ADD_ON_INSTRUCTION GP_HeadPositionDefined   (* revision 1.0 *)
// To be called before invertion data
VAR_IN_OUT
   In_ConvoyData : UDT_Convoy_SL; {required}
END_VAR
VAR_INPUT
   In_dConveyorLenght : DINT; {access None, required}   // Conveyor below [mm/100]
   In_dConveyorWidth : DINT; {access None, required}   // Conveyor below [mm/100]
   In_dInLitePos : DINT; {access None, required}   // Position input lite - Left to Right line flow(0=AX; 1=XA)
   In_dOutDirection : DINT; {required}   // Direction of lateral flow (0=Left; 1=Right; 2=CW(rotation); 3=CCW(rotation))
   In_dOutLitePos : DINT; {access None, required}   // Position output lite - Left to Right line flow(0=AX; 1=XA)
END_VAR
VAR_OUTPUT
   Out_dHeadPosition : DINT; {access Read Only, required}   // New head position [mm/100]
END_VAR
VAR
   TMP_idxCap : DINT; {access None}
   TMP_IdxLite : DINT; {access None}
   TMP_MaxCap : DINT; {access None}
   TMP_MaxLite : DINT; {access None}
   TMP_d : DINT; {access None}
   TMP_LiteHeadReference : DINT; {access None}   // New convoy lite head [mm/100]
END_VAR

ROUTINE Logic   (* structured text *)
   ////////////////////////////////////////////////////////////
   //   Copyright (c)  <Key Automation srl>
   //------------------------------------------------------------
   //   Routine: GP_HeadPositionDefined - Logic
   //   Author: Gerto\admin
   //   Created: 2020-02-05
   //------------------------------------------------------------
   //   Description:
   //
   //
   //   History:
   //
   ////////////////////////////////////////////////////////////
   
   //Dimension array
   Size(In_ConvoyData.rgtCap,0,TMP_MaxCap);
   size(In_ConvoyData.rgtCap[0].rgtLite,0,TMP_MaxLite);
   
   //Find lite of reference
   
   // The smallest LitesHead (Barycenter Lite - 1/2 width lite)
   if 	(In_dOutDirection = 0 and In_dInLitePos = 0 and In_dOutLitePos = 0) or
   	(In_dOutDirection = 0 and In_dInLitePos = 0 and In_dOutLitePos = 1) or
   	(In_dOutDirection = 1 and In_dInLitePos = 1 and In_dOutLitePos = 0) or
   	(In_dOutDirection = 1 and In_dInLitePos = 1 and In_dOutLitePos = 1) or
   	(In_dOutDirection = 2 and In_dInLitePos = 0 and In_dOutLitePos = 0) or
   	(In_dOutDirection = 3 and In_dInLitePos = 1 and In_dOutLitePos = 1) then
   	TMP_LiteHeadReference := In_dConveyorWidth;
   	For TMP_idxCap := 0 to TMP_MaxCap-1 by 1 do
   		for TMP_IdxLite := 0 to TMP_MaxLite-1 by 1 do
   			if In_ConvoyData.rgtCap[TMP_idxCap].rgtLite[TMP_IdxLite].dID <> 0 and (In_ConvoyData.rgtCap[TMP_idxCap].rgtLite[TMP_IdxLite].dBarycenter_cmm - In_ConvoyData.rgtCap[TMP_idxCap].rgtLite[TMP_IdxLite].dWidth_cmm/2) < TMP_LiteHeadReference then
   				TMP_LiteHeadReference := In_ConvoyData.rgtCap[TMP_idxCap].rgtLite[TMP_IdxLite].dBarycenter_cmm - In_ConvoyData.rgtCap[TMP_idxCap].rgtLite[TMP_IdxLite].dWidth_cmm/2;
   			end_if;
   		end_for;
   	end_for;
   end_if;
   
   
   // The biggest LitesHead (Barycenter Lite + 1/2 width lite)
   if 	(In_dOutDirection = 0 and In_dInLitePos = 1 and In_dOutLitePos = 0) or
   	(In_dOutDirection = 0 and In_dInLitePos = 1 and In_dOutLitePos = 1) or
   	(In_dOutDirection = 1 and In_dInLitePos = 0 and In_dOutLitePos = 0) or
   	(In_dOutDirection = 1 and In_dInLitePos = 0 and In_dOutLitePos = 1) or
   	(In_dOutDirection = 2 and In_dInLitePos = 1 and In_dOutLitePos = 1) or
   	(In_dOutDirection = 3 and In_dInLitePos = 0 and In_dOutLitePos = 0) then
   	TMP_LiteHeadReference := 0;
   	For TMP_idxCap := 0 to TMP_MaxCap-1 by 1 do
   		for TMP_IdxLite := 0 to TMP_MaxLite-1 by 1 do
   			if In_ConvoyData.rgtCap[TMP_idxCap].rgtLite[TMP_IdxLite].dID <> 0 and (In_ConvoyData.rgtCap[TMP_idxCap].rgtLite[TMP_IdxLite].dBarycenter_cmm + In_ConvoyData.rgtCap[TMP_idxCap].rgtLite[TMP_IdxLite].dWidth_cmm/2) > TMP_LiteHeadReference then
   				TMP_LiteHeadReference := In_ConvoyData.rgtCap[TMP_idxCap].rgtLite[TMP_IdxLite].dBarycenter_cmm + In_ConvoyData.rgtCap[TMP_idxCap].rgtLite[TMP_IdxLite].dWidth_cmm/2;
   			end_if;
   		end_for;
   	end_for;
   end_if;
   
   //Calculate new head position
   
   // Conveyor deviation
   //Head value = In conveyor width/2 - (barycenter lite - 1/2 lite width) of lite smallest
   if 	(In_dOutDirection = 0 and In_dInLitePos = 0 and In_dOutLitePos = 0) or
   	(In_dOutDirection = 0 and In_dInLitePos = 0 and In_dOutLitePos = 1) or
   	(In_dOutDirection = 1 and In_dInLitePos = 1 and In_dOutLitePos = 0) or
   	(In_dOutDirection = 1 and In_dInLitePos = 1 and In_dOutLitePos = 1) then
   	Out_dHeadPosition := In_dConveyorWidth/2 - TMP_LiteHeadReference;
   end_if;
   
   //Head value = In conveyor width/2 + (barycenter lite + 1/2 lite width) of lite biggest
   if 	(In_dOutDirection = 0 and In_dInLitePos = 1 and In_dOutLitePos = 0) or
   	(In_dOutDirection = 0 and In_dInLitePos = 1 and In_dOutLitePos = 1) or
   	(In_dOutDirection = 1 and In_dInLitePos = 0 and In_dOutLitePos = 0) or
   	(In_dOutDirection = 1 and In_dInLitePos = 0 and In_dOutLitePos = 1) then
   	Out_dHeadPosition := In_dConveyorWidth/2 + TMP_LiteHeadReference;
   end_if;
   
   
   // Rotator
   //Head value = In conveyor lenght / 2 - (baricenter lite - 1/2 lite width) of lite smallest
   if  (In_dOutDirection = 2 and In_dInLitePos = 0 and In_dOutLitePos = 0) or
   	(In_dOutDirection = 3 and In_dInLitePos = 1 and In_dOutLitePos = 1) then
   	Out_dHeadPosition := In_dConveyorLenght/2 - TMP_LiteHeadReference;
   end_if;
   
   // Rotator
   //Head value = In conveyor lenght / 2 + (baricenter lite + 1/2 lite width) of lite biggest
   if  (In_dOutDirection = 2 and In_dInLitePos = 1 and In_dOutLitePos = 1) or
   	(In_dOutDirection = 3 and In_dInLitePos = 0 and In_dOutLitePos = 0) then
   	Out_dHeadPosition := In_dConveyorLenght/2 + TMP_LiteHeadReference;
   end_if;
   
END_ROUTINE
END_ADD_ON_INSTRUCTION

ADD_ON_INSTRUCTION GP_InvertCapxLite   (* revision 1.0 *)
VAR_INPUT
   In_dInLitePos : DINT; {access None, required}   // Position input lite - Left to Right line flow(0=AX; 1=XA)
   In_dOutLitePos : DINT; {access None, required}   // Position output lite - Left to Right line flow(0=AX; 1=XA)
   In_dOutDirection : DINT; {required}   // Direction of lateral flow (0=Left; 1=Right; 2=CW(rotation); 3=CCW(rotation))
END_VAR
VAR_IN_OUT
   In_ConvoyData : UDT_Convoy_SL; {required}
   Out_ConvoyData : UDT_Convoy_SL; {required}
   Const_ConvoyData_Empty : UDT_Convoy_SL; {constant, required}
END_VAR
VAR_INPUT
   In_dConveyorLength : DINT; {access None, required}   // Conveyor below [mm/100]
   In_dConveyorWidth : DINT; {access None, required}   // Conveyor below [mm/100]
END_VAR
VAR_OUTPUT
   Out_dHeadPosition : DINT; {access Read Only, required}   // New head position [mm/100]
END_VAR
VAR_INPUT
   In_dHeadPosition : DINT; {required}   // Head position on conveyor below [mm/100]
   In_dOffset1 : DINT; {required}   // Distance of start conveyorIn and axe conveyorOut [mm/100]
   In_dOffset2 : DINT;   // Distance between stop conveyorOut and stop conveyorIn [mm/100] (NU)
END_VAR
VAR_OUTPUT
   Out_dCause : DINT; {access Read Only}
END_VAR
VAR
   TMP_MaxCapIn : DINT; {access None}
   TMP_MaxLiteIn : DINT; {access None}
   TMP_idxInCap : DINT; {access None}
   TMP_IdxInLite : DINT; {access None}
   TMP_MaxCapOut : DINT; {access None}
   TMP_MaxLiteOut : DINT; {access None}
   TMP_IdxOutCap : DINT; {access None}
   TMP_IdxOutLite : DINT; {access None}
   TMP_d : DINT; {access None}
   GP_CompactConvoy : GP_CompactConvoy; {access None}
   GP_HeadPositionDefined : GP_HeadPositionDefined; {access None}
   GP_BaricenterDefinition : GP_BaricenterDefinition; {access None}
   TMP_In_ConvoyData : UDT_Convoy_SL; {access None}
   TMP_Idx : DINT; {access None}
   TMP_YPosMinus : DINT[10]; {access None}
   TMP_YPosPlus : DINT[10]; {access None}
   TMP_nNoLiteFound : DINT; {access None}
   TMP_Idx2 : DINT; {access None}
   GP_CompactConvoy_V2 : GP_CompactConvoy_V2; {access None}
END_VAR

ROUTINE Logic   (* structured text *)
   ////////////////////////////////////////////////////////////
   //   Copyright (c)  <Key Automation srl>
   //------------------------------------------------------------
   //   Routine: GP_InvertCapxLite - Logic
   //   Author: Gerto
   //   Created: 2020-02-03
   //------------------------------------------------------------
   //   Description:
   //
   //
   //   History:
   //
   ////////////////////////////////////////////////////////////
   
   cop(In_ConvoyData,TMP_In_ConvoyData,1);
   
   //Dimension array
   Size(In_ConvoyData.rgtCap,0,TMP_MaxCapIn);
   size(TMP_In_ConvoyData.rgtCap[0].rgtLite,0,TMP_MaxLiteIn);
   Size(Out_ConvoyData.rgtCap,0,TMP_MaxCapOut);
   size(Out_ConvoyData.rgtCap[0].rgtLite,0,TMP_MaxLiteOut);
   
   //Init
   cop(Const_ConvoyData_Empty,Out_ConvoyData,1);
   TMP_nNoLiteFound := -999999999;
   Out_dCause := 0;
   
   
   //Definition Head position (before rotation data CapxLite)
   GP_HeadPositionDefined(GP_HeadPositionDefined,TMP_In_ConvoyData,In_dConveyorLength,In_dConveyorWidth,In_dInLitePos,In_dOutDirection,In_dOutLitePos,Out_dHeadPosition);
   
   //Definition baricenter (before rotation data CapxLite)
   GP_BaricenterDefinition(GP_BaricenterDefinition,In_dHeadPosition,TMP_In_ConvoyData,In_dInLitePos,In_dOutDirection,In_dOutLitePos,In_dOffset1,In_dOffset2,In_dConveyorLength,In_dConveyorWidth);
   
   
   
   // Input cap //////////////////////////////////////////////////
   //
   For TMP_idxInCap := TMP_In_ConvoyData.dTotalCaps-1 to 0 by -1 do
   
   	if 	(In_dOutDirection = 0 and In_dInLitePos = 0 and In_dOutLitePos = 0) or
   		(In_dOutDirection = 0 and In_dInLitePos = 1 and In_dOutLitePos = 0) or
   		(In_dOutDirection = 1 and In_dInLitePos = 0 and In_dOutLitePos = 1) or
   		(In_dOutDirection = 1 and In_dInLitePos = 1 and In_dOutLitePos = 1) or
   		(In_dOutDirection = 2 and In_dInLitePos = 0 and In_dOutLitePos = 0) or
   		(In_dOutDirection = 3 and In_dInLitePos = 1 and In_dOutLitePos = 1) then
   			TMP_IdxOutLite :=  TMP_In_ConvoyData.dTotalCaps-1 - TMP_idxInCap;		// last cap to first lite
   	end_if;
   
   	if 	(In_dOutDirection = 0 and In_dInLitePos = 0 and In_dOutLitePos = 1) or
   		(In_dOutDirection = 0 and In_dInLitePos = 1 and In_dOutLitePos = 1) or
   		(In_dOutDirection = 1 and In_dInLitePos = 0 and In_dOutLitePos = 0) or
   		(In_dOutDirection = 1 and In_dInLitePos = 1 and In_dOutLitePos = 0) or
   		(In_dOutDirection = 2 and In_dInLitePos = 1 and In_dOutLitePos = 1) or
   		(In_dOutDirection = 3 and In_dInLitePos = 0 and In_dOutLitePos = 0) then
   			TMP_IdxOutLite := TMP_idxInCap;										// last cap to last lite
   	end_if;
   
   	For TMP_IdxInLite := TMP_MaxLiteIn-1 to 0 by -1 do
   
   		if 	(In_dOutDirection = 0 and In_dInLitePos = 1 and In_dOutLitePos = 0) or
   			(In_dOutDirection = 0 and In_dInLitePos = 1 and In_dOutLitePos = 1) or
   			(In_dOutDirection = 1 and In_dInLitePos = 0 and In_dOutLitePos = 0) or
   			(In_dOutDirection = 1 and In_dInLitePos = 0 and In_dOutLitePos = 1) or
   			(In_dOutDirection = 2 and In_dInLitePos = 1 and In_dOutLitePos = 1) or
   			(In_dOutDirection = 3 and In_dInLitePos = 0 and In_dOutLitePos = 0) then
   				TMP_IdxOutCap := TMP_MaxLiteIn-1 - TMP_IdxInLite;			// last lite to first cap
   		end_if;
   
   		if 	(In_dOutDirection = 0 and In_dInLitePos = 0 and In_dOutLitePos = 0) or
   			(In_dOutDirection = 0 and In_dInLitePos = 0 and In_dOutLitePos = 1) or
   			(In_dOutDirection = 1 and In_dInLitePos = 1 and In_dOutLitePos = 0) or
   			(In_dOutDirection = 1 and In_dInLitePos = 1 and In_dOutLitePos = 1) or
   			(In_dOutDirection = 2 and In_dInLitePos = 0 and In_dOutLitePos = 0) or
   			(In_dOutDirection = 3 and In_dInLitePos = 1 and In_dOutLitePos = 1) then
   				TMP_IdxOutCap := TMP_IdxInLite;									// last lite to last cap
   		end_if;
   		// copy data lite
   		if TMP_In_ConvoyData.rgtCap[TMP_idxInCap].rgtLite[TMP_IdxInLite].dID <> 0 then
   			cop(TMP_In_ConvoyData.rgtCap[TMP_idxInCap].rgtLite[TMP_IdxInLite],Out_ConvoyData.rgtCap[TMP_IdxOutCap].rgtLite[TMP_IdxOutLite],1);
   		end_if;
   		//Write cap length from lite width
   		if TMP_In_ConvoyData.rgtCap[TMP_idxInCap].rgtLite[TMP_IdxInLite].dWidth_cmm > 0 then
   			Out_ConvoyData.rgtCap[TMP_IdxOutCap].dLength_cmm := TMP_In_ConvoyData.rgtCap[TMP_idxInCap].rgtLite[TMP_IdxInLite].dWidth_cmm;
   		end_if;
   
   		// Write lite width from cap length
   		if Out_ConvoyData.rgtCap[TMP_IdxOutCap].rgtLite[TMP_IdxOutLite].dID <>0 then
   			Out_ConvoyData.rgtCap[TMP_IdxOutCap].rgtLite[TMP_IdxOutLite].dWidth_cmm := TMP_In_ConvoyData.rgtCap[TMP_idxInCap].dLength_cmm;
   		end_if;
   	end_for;
   end_for;
   
   //gap between cap (calculate with in_baricenter lite difference)
   //init Y position
   for TMP_Idx := 0 to 10-1 by 1 do
   	TMP_YPosMinus[TMP_Idx] := 0;
   	TMP_YPosPlus[TMP_Idx] := 0;
   end_for;
   	//save Y position value
   for TMP_IdxInLite := 0 to TMP_MaxLiteIn-1 by 1 do
   	for TMP_idxInCap := 0 to TMP_MaxCapIn-1 by 1 do
   		if TMP_In_ConvoyData.rgtCap[TMP_idxInCap].rgtLite[TMP_IdxInLite].dID <> 0 then
   			TMP_YPosMinus[TMP_IdxInLite] := In_ConvoyData.rgtCap[TMP_idxInCap].rgtLite[TMP_IdxInLite].dBarycenter_cmm - In_ConvoyData.rgtCap[TMP_idxInCap].rgtLite[TMP_IdxInLite].dWidth_cmm / 2;
   			TMP_YPosPlus[TMP_IdxInLite] := In_ConvoyData.rgtCap[TMP_idxInCap].rgtLite[TMP_IdxInLite].dBarycenter_cmm + In_ConvoyData.rgtCap[TMP_idxInCap].rgtLite[TMP_IdxInLite].dWidth_cmm / 2;
   			exit;
   		else; //no lite found
   			TMP_YPosMinus[TMP_IdxInLite] := TMP_nNoLiteFound;
   			TMP_YPosPlus[TMP_IdxInLite] := TMP_nNoLiteFound;
   		end_if;
   	end_for;
   end_for;
   	//write data gap to output gap
   for TMP_IdxOutCap := 0 to TMP_MaxCapOut-1 by 1  do
   	if 	(In_dOutDirection = 0 and In_dInLitePos = 0 and In_dOutLitePos = 0) or
   		(In_dOutDirection = 0 and In_dInLitePos = 0 and In_dOutLitePos = 1) or
   		(In_dOutDirection = 1 and In_dInLitePos = 1 and In_dOutLitePos = 0) or
   		(In_dOutDirection = 1 and In_dInLitePos = 1 and In_dOutLitePos = 1) or
   		(In_dOutDirection = 2 and In_dInLitePos = 0 and In_dOutLitePos = 0) or
   		(In_dOutDirection = 3 and In_dInLitePos = 1 and In_dOutLitePos = 1) then //first lite in first cap out
   		TMP_Idx := TMP_IdxOutCap;
   	end_if;
   	if 	(In_dOutDirection = 0 and In_dInLitePos = 1 and In_dOutLitePos = 0) or
   		(In_dOutDirection = 0 and In_dInLitePos = 1 and In_dOutLitePos = 1) or
   		(In_dOutDirection = 1 and In_dInLitePos = 0 and In_dOutLitePos = 0) or
   		(In_dOutDirection = 1 and In_dInLitePos = 0 and In_dOutLitePos = 1) or
   		(In_dOutDirection = 2 and In_dInLitePos = 1 and In_dOutLitePos = 1) or
   		(In_dOutDirection = 3 and In_dInLitePos = 0 and In_dOutLitePos = 0) then //first lite in last cap out
   		TMP_Idx := TMP_MaxCapOut -1 - TMP_IdxOutCap;
   	end_if;
   
   	//find first TMP_YPosMinus[TMP_Idx+1] <> TMP_nNoLiteFound
   	for TMP_Idx2 := TMP_Idx+1 to 10-1 by 1 do
   		if TMP_YPosMinus[TMP_Idx2] <> TMP_nNoLiteFound then
   			TMP_d := TMP_YPosMinus[TMP_Idx2];
   			exit;
   		else;
   		TMP_d := TMP_nNoLiteFound;
   		end_if;
   	end_for;
   	// if tMP_d <> TMP_nNoLiteFound (lite found) calculate gap
   	if TMP_d <> TMP_nNoLiteFound and TMP_YPosPlus[TMP_Idx] <> TMP_nNoLiteFound then
   	Out_ConvoyData.rgtCap[TMP_IdxOutCap].dReqGapForConv_cmm := TMP_d - TMP_YPosPlus[TMP_Idx];
   	end_if;
   	if Out_ConvoyData.rgtCap[TMP_IdxOutCap].dReqGapForConv_cmm < 0 then
   		Out_ConvoyData.rgtCap[TMP_IdxOutCap].dReqGapForConv_cmm := 0;
   		Out_dCause := 100; //gap finded < 0
   	end_if;
   end_for;
   
   //Data convoy
   //Convoy length calculated in "compact convoy"
   Out_ConvoyData.dGapCaps_cmm	:= TMP_In_ConvoyData.rgtCap[0].dGap_cmm; //gap between caps
   
   ////Data Caps
   //for TMP_IdxOutCap := 0 to TMP_In_ConvoyData.rgtCap[0].dNumLites - 1 by 1 do
   //	Out_ConvoyData.rgtCap[TMP_IdxOutCap].dNumLites := TMP_In_ConvoyData.dTotalCaps; 					//qta lite
   //	if Out_ConvoyData.rgtCap[TMP_IdxOutCap].dNumLites < 1 then
   //		Out_ConvoyData.rgtCap[TMP_IdxOutCap].dNumLites := 1;
   //	end_if;
   //	Out_ConvoyData.rgtCap[TMP_IdxOutCap].dGap_cmm := TMP_In_ConvoyData.dGapCaps_cmm;					//gaps between lites
   //	Out_ConvoyData.rgtCap[TMP_IdxOutCap].dWidth_cmm := TMP_In_ConvoyData.dLength_cmm;					//total cap(convoy) width
   //	Out_ConvoyData.rgtCap[TMP_IdxOutCap].dThickness_cmm := TMP_In_ConvoyData.rgtCap[0].dThickness_cmm;	//thikness cap
   //end_for;
   ////Write capID (first LiteID finded)
   //For TMP_IdxOutCap := 0 to TMP_MaxCapOut-1 by 1 do
   //	For TMP_IdxOutLite := 0 to TMP_MaxLiteOut-1 by 1 do
   //		if Out_ConvoyData.rgtCap[TMP_IdxOutCap].rgtLite[TMP_IdxOutLite].dID <>0 then
   //			Out_ConvoyData.rgtCap[TMP_IdxOutCap].dID := Out_ConvoyData.rgtCap[TMP_IdxOutCap].rgtLite[TMP_IdxOutLite].dID;
   //			exit;
   //		end_if;
   //	end_for;
   //end_for;
   
   FOR TMP_IdxOutCap := 0 TO TMP_MaxCapOut - 1 BY 1 DO
       FOR TMP_IdxOutLite := 0 TO TMP_MaxLiteOut - 1 BY 1 DO
           IF Out_ConvoyData.rgtCap[TMP_IdxOutCap].rgtLite[TMP_IdxOutLite].dID <> 0 THEN
               Out_ConvoyData.rgtCap[TMP_IdxOutCap].dID := Out_ConvoyData.rgtCap[TMP_IdxOutCap].rgtLite[TMP_IdxOutLite].dID;
               Out_ConvoyData.rgtCap[TMP_IdxOutCap].dNumLites := TMP_In_ConvoyData.dTotalCaps;                     //qta lite
               IF Out_ConvoyData.rgtCap[TMP_IdxOutCap].dNumLites < 1 THEN
                   Out_ConvoyData.rgtCap[TMP_IdxOutCap].dNumLites := 1;
               END_IF;
               Out_ConvoyData.rgtCap[TMP_IdxOutCap].dWidth_cmm := TMP_In_ConvoyData.dLength_cmm;                   //total cap(convoy) width
               Out_ConvoyData.rgtCap[TMP_IdxOutCap].dThickness_cmm := TMP_In_ConvoyData.rgtCap[0].dThickness_cmm;  //thikness cap
               EXIT;
           END_IF;
       END_FOR;
   END_FOR;
   
   //Compact convoy
   GP_CompactConvoy(GP_CompactConvoy,Out_ConvoyData,Const_ConvoyData_Empty);
   
END_ROUTINE
END_ADD_ON_INSTRUCTION

ADD_ON_INSTRUCTION GP_NetworkDiag   (* revision 1.0 *)
VAR_IN_OUT
   IN_OB_Initialize : GP_OB_Initialize; {required}
   IN_ModuleName : MODULE; {required}   // Module name
   OUT_tModuleInfo : GP_NetworkDiag_v1; {required}   // Module info
END_VAR
VAR
   TMP_xFaulted : BOOL; {access None}
   TMP_xConnected : BOOL; {access None}
END_VAR

ROUTINE Logic   (* structured text *)
   //Initialize
   TMP_xConnected:=0;
   TMP_xFaulted:=0;
   
   //Get system info from module
   gsv(Module,IN_ModuleName,EntryStatus,OUT_tModuleInfo.dEntryStatus);
   gsv(Module,IN_ModuleName,FaultCode,OUT_tModuleInfo.dFaultCode);
   gsv(Module,IN_ModuleName,FaultInfo,OUT_tModuleInfo.dFaultInfo);
   gsv(Module,IN_ModuleName,Instance,OUT_tModuleInfo.dInstance);
   
   CASE OUT_tModuleInfo.dEntryStatus OF
   	16#0000:(*Standby: the controller is powering up.*)
    			TMP_xFaulted:= IN_OB_Initialize.OUT_xClock_800ms;
   
   	16#1000:(*Faulted: any of the MODULE object’s connections to the associated module fail.
   			This value should not be used to determine if the module failed because the MODULE
   			object leaves this state periodically when trying to reconnect to the module.
   			Instead, test for Running state (164000). Check for FaultCode not equal to 0 to determine if a module is faulted.
   			When Faulted, the FaultCode and FaultInfo attributes are valid until the fault condition is corrected.*)
    			TMP_xConnected:= IN_OB_Initialize.OUT_xClock_1s;
   			TMP_xFaulted:= 1;
   
   	16#2000:(*Validating: the MODULE object is verifying MODULE object integrity prior to establishing connections to the module.*)
    			TMP_xConnected:= IN_OB_Initialize.OUT_xClock_400ms;
   
   	16#3000:(*Connecting: the MODULE object is initiating connections to the module.*)
   			TMP_xConnected:= IN_OB_Initialize.OUT_xClock_400ms;
   
   	16#4000:(*Running: all connections to the module are established and data is successfully transferring.*)
    			TMP_xConnected:= 1;
   
   	16#5000:(*Shutting down: the MODULE object is in the process of shutting down all connections to the module.*)
   			TMP_xConnected:= IN_OB_Initialize.OUT_xClock_1s;
   
   	16#6000:(*Inhibited: the MODULE object is inhibited (the inhibit bit in the Mode attribute is set).*)
    			TMP_xConnected:= IN_OB_Initialize.OUT_xClock_1s;
   
   	16#7000:(*Waiting: the parent MODULE object upon which this MODULE object depends is not running*)
   			TMP_xConnected:= IN_OB_Initialize.OUT_xClock_1s;
   
   	16#9000:(*FirmwareUpdating: Firmware supervisor is attempting to flash the module. *)
    			TMP_xConnected:= IN_OB_Initialize.OUT_xClock_800ms;
   
   	16#A000:(*Configuring: Controller is downloading configuration to the module.
   			Either ?forward open? or (ADC) download occur during this state.*)
   			TMP_xConnected:= IN_OB_Initialize.OUT_xClock_800ms;
   END_CASE;
   
   IF OUT_tModuleInfo.dFaultCode<>0 THEN
   	TMP_xFaulted:= 1;
   END_IF;
   
   //Save status bit
   OUT_tModuleInfo.xConnected:=TMP_xConnected;
   OUT_tModuleInfo.xFaulted:=TMP_xFaulted;
   
   
   
   
   
   
   
   
   
   
   
   
   
   
   
   
   
   
   
   
END_ROUTINE
END_ADD_ON_INSTRUCTION

ADD_ON_INSTRUCTION GP_OB_Initialize   (* revision 1.0 *)
VAR_IN_OUT
   STC : GP_OB_Initialize_STC; {required}
END_VAR
VAR_INPUT
   IN_xInitialize : BOOL; {access None, required}   // Initialize values (Restart call)
END_VAR
VAR_OUTPUT
   OUT_dExecutionTime_ms : DINT; {access None}   // OB Execution time [ms]
   OUT_dMinExecutionTime_ms : DINT; {access None}   // OB Minimum execution time [ms]
   OUT_dMaxExecutionTime_ms : DINT; {access None}   // OB Maximum execution time [ms]
   OUT_xOs_100ms : BOOL; {access None}   // OS each 100ms
   OUT_xOs_200ms : BOOL; {access None}   // OS each 200ms
   OUT_xOs_400ms : BOOL; {access None}   // OS each 400ms
   OUT_xOs_500ms : BOOL; {access None}   // OS each 500ms
   OUT_xOs_800ms : BOOL; {access None}   // OS each 800ms
   OUT_xOs_1s : BOOL; {access None}   // OS each 1s
   OUT_xOs_2s : BOOL; {access None}   // OS each 2s
   OUT_xOs_5s : BOOL; {access None}   // OS each 5s
   OUT_xOs_10s : BOOL; {access None}   // OS each 10s
   OUT_xOs_30s : BOOL; {access None}   // OS each 30s
   OUT_xOs_1min : BOOL; {access None}   // OS each 1min
   OUT_xOs_2min : BOOL; {access None}   // OS each 2min
   OUT_xOs_10min : BOOL; {access None}   // OS each 10min
   OUT_xOs_30min : BOOL; {access None}   // OS each 30min
   OUT_xOs_1h : BOOL; {access None}   // OS each 1h
   OUT_xClock_100ms : BOOL; {access None}   // Clock 100ms
   OUT_xClock_200ms : BOOL; {access None}   // Clock 200ms
   OUT_xClock_400ms : BOOL; {access None}   // Clock 400ms
   OUT_xClock_500ms : BOOL; {access None}   // Clock 500ms
   OUT_xClock_800ms : BOOL; {access None}   // Clock 800ms
   OUT_xClock_1s : BOOL; {access None}   // Clock 1s
   OUT_xClock_2s : BOOL; {access None}   // Clock 2s
   OUT_xClock_5s : BOOL; {access None}   // Clock 5s
   OUT_xClock_10s : BOOL; {access None}   // Clock 10s
   OUT_xClock_30s : BOOL; {access None}   // Clock 30s
   OUT_xClock_1min : BOOL; {access None}   // Clock 1min
   OUT_xClock_2min : BOOL; {access None}   // Clock 2min
   OUT_xClock_10min : BOOL; {access None}   // Clock 10min
   OUT_xClock_30min : BOOL; {access None}   // Clock 30min
   OUT_xClock_1h : BOOL; {access None}   // Clock 1h
   OUT_xDebugOFF : BOOL; {access None}
   OUT_xDebugON : BOOL; {access None}
END_VAR
VAR
   CONST_DMAX_INT : DINT; {access None}
   CONST_DTICK_1H : DINT; {access None}
   CONST_DTICK_30MIN : DINT; {access None}
   CONST_DTICK_10MIN : DINT; {access None}
   CONST_DTICK_2MIN : DINT; {access None}
   CONST_DTICK_1MIN : DINT; {access None}
   CONST_DTICK_30S : DINT; {access None}
   CONST_DTICK_10S : DINT; {access None}
   CONST_DTICK_5S : DINT; {access None}
   CONST_DTICK_2S : DINT; {access None}
   CONST_DTICK_1S : DINT; {access None}
   CONST_DTICK_800MS : DINT; {access None}
   CONST_DTICK_500MS : DINT; {access None}
   CONST_DTICK_400MS : DINT; {access None}
   CONST_DTICK_200MS : DINT; {access None}
   CONST_DTICK_100MS : DINT; {access None}
   TMP_rlActualExecutionTimeRound : REAL; {access None}   // Rounded execution time [ms]
   TMP_rlActualExecutionTime : REAL; {access None}   // ActualExecutionTime [ms]
END_VAR

ROUTINE Logic   (* structured text *)
   //Costants
   CONST_DTICK_100MS:=100;
   CONST_DTICK_200MS:=200;
   CONST_DTICK_400MS:=400;
   CONST_DTICK_500MS:=500;
   CONST_DTICK_800MS:=800;
   CONST_DTICK_1S:=1000;
   CONST_DTICK_2S:=2000;
   CONST_DTICK_5S:=5000;
   CONST_DTICK_10S:=10000;
   CONST_DTICK_30S:=30000;
   CONST_DTICK_1MIN:=60000;
   CONST_DTICK_2MIN:=120000;
   CONST_DTICK_10MIN:=600000;
   CONST_DTICK_30MIN:=1800000;
   CONST_DTICK_1H:=86400000;
   CONST_DMAX_INT:=16#7FFFFFFF;
   OUT_xDebugOFF:=0;
   OUT_xDebugON:=1;
   
   //Initialize OS bits
   OUT_xOs_100ms := 0;
   OUT_xOs_200ms := 0;
   OUT_xOs_400ms := 0;
   OUT_xOs_500ms := 0;
   OUT_xOs_800ms := 0;
   OUT_xOs_1s := 0;
   OUT_xOs_2s := 0;
   OUT_xOs_5s := 0;
   OUT_xOs_10s := 0;
   OUT_xOs_30s := 0;
   OUT_xOs_1min := 0;
   OUT_xOs_2min := 0;
   OUT_xOs_10min := 0;
   OUT_xOs_30min := 0;
   OUT_xOs_1h := 0;
   
   //Take the start execution time from the CPU
   gsv(Task,THIS,StartTime,STC.lwStartTime[0]);
   
   //Initialize FB execution
   IF IN_xInitialize THEN
   
   	IN_xInitialize := 0;
   	OUT_dExecutionTime_ms := 0;
   	OUT_dMinExecutionTime_ms := CONST_DMAX_INT;
   	OUT_dMaxExecutionTime_ms := 0;
   	OUT_xClock_100ms := 0;
   	OUT_xClock_200ms := 0;
   	OUT_xClock_400ms := 0;
   	OUT_xClock_500ms := 0;
   	OUT_xClock_800ms := 0;
   	OUT_xClock_1s := 0;
   	OUT_xClock_2s := 0;
   	OUT_xClock_5s := 0;
   	OUT_xClock_10s := 0;
   	OUT_xClock_30s := 0;
   	OUT_xClock_1min := 0;
   	OUT_xClock_2min := 0;
   	OUT_xClock_10min := 0;
   	OUT_xClock_30min := 0;
   	OUT_xClock_1h := 0;
   
   	STC.dElapsed_100ms_ms := 0;
   	STC.dElapsed_200ms_ms := 0;
   	STC.dElapsed_400ms_ms := 0;
   	STC.dElapsed_500ms_ms := 0;
   	STC.dElapsed_800ms_ms := 0;
   	STC.dElapsed_1s_ms := 0;
   	STC.dElapsed_2s_ms := 0;
   	STC.dElapsed_5s_ms := 0;
   	STC.dElapsed_10s_ms := 0;
   	STC.dElapsed_30s_ms := 0;
   	STC.dElapsed_1min_ms := 0;
   	STC.dElapsed_2min_ms := 0;
   	STC.dElapsed_10min_ms := 0;
   	STC.dElapsed_30min_ms := 0;
   	STC.dElapsed_1h_ms := 0;
   
   	STC.lwOldStartTime[0] := STC.lwStartTime[0];
   	STC.lwOldStartTime[1] := STC.lwStartTime[1];
   
   END_IF;
   
   //***** CALCULATE OB EXECUTION TIME *****
   STC.dlLastExecValue_us := STC.lwStartTime[0] - STC.lwOldStartTime[0];
   STC.lwOldStartTime[0] := STC.lwStartTime[0];
   STC.lwOldStartTime[1] := STC.lwStartTime[1];
   //Convert from [us] to [ms]
   TMP_rlActualExecutionTime := STC.dlLastExecValue_us / 1000.0;
   //Add the reminder of the last cycle
   TMP_rlActualExecutionTime := TMP_rlActualExecutionTime + STC.rReminder_ms;
   //Calculate the rounded value
   TMP_rlActualExecutionTimeRound:= trunc(TMP_rlActualExecutionTime + 0.5);
   OUT_dExecutionTime_ms := trunc(TMP_rlActualExecutionTime + 0.5);
   //Save the reminder for the next cycle
   STC.rReminder_ms := TMP_rlActualExecutionTime - TMP_rlActualExecutionTimeRound;
   
   //Save the maximum scan value
   IF OUT_dExecutionTime_ms > OUT_dMaxExecutionTime_ms THEN
   	OUT_dMaxExecutionTime_ms := OUT_dExecutionTime_ms;
   END_IF;
   
   //Save the minimum scan value
   IF OUT_dExecutionTime_ms < OUT_dMinExecutionTime_ms THEN
   	OUT_dMinExecutionTime_ms := OUT_dExecutionTime_ms;
   END_IF;
   
   //***** CALCULATE SERVICES CLOCK *****
   
   //Increment counters for each clock
   STC.dElapsed_100ms_ms := STC.dElapsed_100ms_ms + OUT_dExecutionTime_ms;
   STC.dElapsed_200ms_ms := STC.dElapsed_200ms_ms + OUT_dExecutionTime_ms;
   STC.dElapsed_400ms_ms := STC.dElapsed_400ms_ms + OUT_dExecutionTime_ms;
   STC.dElapsed_500ms_ms := STC.dElapsed_500ms_ms + OUT_dExecutionTime_ms;
   STC.dElapsed_800ms_ms := STC.dElapsed_800ms_ms + OUT_dExecutionTime_ms;
   STC.dElapsed_1s_ms := STC.dElapsed_1s_ms + OUT_dExecutionTime_ms;
   STC.dElapsed_2s_ms := STC.dElapsed_2s_ms + OUT_dExecutionTime_ms;
   STC.dElapsed_5s_ms := STC.dElapsed_5s_ms + OUT_dExecutionTime_ms;
   STC.dElapsed_10s_ms := STC.dElapsed_10s_ms + OUT_dExecutionTime_ms;
   STC.dElapsed_30s_ms := STC.dElapsed_30s_ms + OUT_dExecutionTime_ms;
   STC.dElapsed_1min_ms := STC.dElapsed_1min_ms + OUT_dExecutionTime_ms;
   STC.dElapsed_2min_ms := STC.dElapsed_2min_ms + OUT_dExecutionTime_ms;
   STC.dElapsed_10min_ms := STC.dElapsed_10min_ms + OUT_dExecutionTime_ms;
   STC.dElapsed_30min_ms := STC.dElapsed_30min_ms + OUT_dExecutionTime_ms;
   STC.dElapsed_1h_ms := STC.dElapsed_1h_ms + OUT_dExecutionTime_ms;
   
   //Calculate the 100ms
   IF STC.dElapsed_100ms_ms >= CONST_DTICK_100MS THEN
   	STC.dElapsed_100ms_ms := STC.dElapsed_100ms_ms - CONST_DTICK_100MS;
   
   	OUT_xOs_100ms := 1;
   
   	IF NOT(OUT_xClock_100ms) THEN
   		OUT_xClock_100ms := 1;
   	ELSE
   		OUT_xClock_100ms := 0;
   	END_IF;
   END_IF;
   
   //Calculate the 200ms
   IF STC.dElapsed_200ms_ms >= CONST_DTICK_200MS THEN
   	STC.dElapsed_200ms_ms := STC.dElapsed_200ms_ms - CONST_DTICK_200MS;
   
   	OUT_xOs_200ms := 1;
   
   	IF NOT(OUT_xClock_200ms) THEN
   		OUT_xClock_200ms := 1;
   	ELSE
   		OUT_xClock_200ms := 0;
   	END_IF;
   END_IF;
   
   //Calculate the 400ms
   IF STC.dElapsed_400ms_ms >= CONST_DTICK_400MS THEN
   	STC.dElapsed_400ms_ms := STC.dElapsed_400ms_ms - CONST_DTICK_400MS;
   
   	OUT_xOs_400ms := 1;
   
   	IF NOT(OUT_xClock_400ms) THEN
   		OUT_xClock_400ms := 1;
   	ELSE
   		OUT_xClock_400ms := 0;
   	END_IF;
   END_IF;
   
   //Calculate the 500ms
   IF STC.dElapsed_500ms_ms >= CONST_DTICK_500MS THEN
   	STC.dElapsed_500ms_ms := STC.dElapsed_500ms_ms - CONST_DTICK_500MS;
   
   	OUT_xOs_500ms := 1;
   
   	IF NOT(OUT_xClock_500ms) THEN
   		OUT_xClock_500ms := 1;
   	ELSE
   		OUT_xClock_500ms := 0;
   	END_IF;
   END_IF;
   
   //Calculate the 800ms
   IF STC.dElapsed_800ms_ms >= CONST_DTICK_800MS THEN
   	STC.dElapsed_800ms_ms := STC.dElapsed_800ms_ms - CONST_DTICK_800MS;
   
   	OUT_xOs_800ms := 1;
   
   	IF NOT(OUT_xClock_800ms) THEN
   		OUT_xClock_800ms := 1;
   	ELSE
   		OUT_xClock_800ms := 0;
   	END_IF;
   END_IF;
   
   //Calculate the 1s
   IF STC.dElapsed_1s_ms >= CONST_DTICK_1S THEN
   	STC.dElapsed_1s_ms := STC.dElapsed_1s_ms - CONST_DTICK_1S;
   
   	OUT_xOs_1s := 1;
   
   	IF NOT(OUT_xClock_1s) THEN
   		OUT_xClock_1s := 1;
   	ELSE
   		OUT_xClock_1s := 0;
   	END_IF;
   END_IF;
   
   //Calculate the 2s
   IF STC.dElapsed_2s_ms >= CONST_DTICK_2S THEN
   	STC.dElapsed_2s_ms := STC.dElapsed_2s_ms - CONST_DTICK_2S;
   
   	OUT_xOs_2s := 1;
   
   	IF NOT(OUT_xClock_2s) THEN
   		OUT_xClock_2s := 1;
   	ELSE
   		OUT_xClock_2s := 0;
   	END_IF;
   END_IF;
   
   //Calculate the 5s
   IF STC.dElapsed_5s_ms >= CONST_DTICK_5S THEN
   	STC.dElapsed_5s_ms := STC.dElapsed_5s_ms - CONST_DTICK_5S;
   
   	OUT_xOs_5s := 1;
   
   	IF NOT(OUT_xClock_5s) THEN
   		OUT_xClock_5s := 1;
   	ELSE
   		OUT_xClock_5s := 0;
   	END_IF;
   END_IF;
   
   //Calculate the 10s
   IF STC.dElapsed_10s_ms >= CONST_DTICK_10S THEN
   	STC.dElapsed_10s_ms := STC.dElapsed_10s_ms - CONST_DTICK_10S;
   
   	OUT_xOs_10s := 1;
   
   	IF NOT(OUT_xClock_10s) THEN
   		OUT_xClock_10s := 1;
   	ELSE
   		OUT_xClock_10s := 0;
   	END_IF;
   END_IF;
   
   //Calculate the 30s
   IF STC.dElapsed_30s_ms >= CONST_DTICK_30S THEN
   	STC.dElapsed_30s_ms := STC.dElapsed_30s_ms - CONST_DTICK_30S;
   
   	OUT_xOs_30s := 1;
   
   	IF NOT(OUT_xClock_30s) THEN
   		OUT_xClock_30s := 1;
   	ELSE
   		OUT_xClock_30s := 0;
   	END_IF;
   END_IF;
   
   //Calculate the 1min
   IF STC.dElapsed_1min_ms >= CONST_DTICK_1MIN THEN
   	STC.dElapsed_1min_ms := STC.dElapsed_1min_ms - CONST_DTICK_1MIN;
   
   	OUT_xOs_1min := 1;
   
   	IF NOT(OUT_xClock_1min) THEN
   		OUT_xClock_1min := 1;
   	ELSE
   		OUT_xClock_1min := 0;
   	END_IF;
   END_IF;
   
   //Calculate the 2min
   IF STC.dElapsed_2min_ms >= CONST_DTICK_2MIN THEN
   	STC.dElapsed_2min_ms := STC.dElapsed_2min_ms - CONST_DTICK_2MIN;
   
   	OUT_xOs_2min := 1;
   
   	IF NOT(OUT_xClock_2min) THEN
   		OUT_xClock_2min := 1;
   	ELSE
   		OUT_xClock_2min := 0;
   	END_IF;
   END_IF;
   
   //Calculate the 10min
   IF STC.dElapsed_10min_ms >= CONST_DTICK_10MIN THEN
   	STC.dElapsed_10min_ms := STC.dElapsed_10min_ms - CONST_DTICK_10MIN;
   
   	OUT_xOs_10min := 1;
   
   	IF NOT(OUT_xClock_10min) THEN
   		OUT_xClock_10min := 1;
   	ELSE
   		OUT_xClock_10min := 0;
   	END_IF;
   END_IF;
   
   //Calculate the 30min
   IF STC.dElapsed_30min_ms >= CONST_DTICK_30MIN THEN
   	STC.dElapsed_30min_ms := STC.dElapsed_30min_ms - CONST_DTICK_30MIN;
   
   	OUT_xOs_30min := 1;
   
   	IF NOT(OUT_xClock_30min) THEN
   		OUT_xClock_30min := 1;
   	ELSE
   		OUT_xClock_30min := 0;
   	END_IF;
   END_IF;
   
   //Calculate the 1h
   IF STC.dElapsed_1h_ms >= CONST_DTICK_1H THEN
   	STC.dElapsed_1h_ms := STC.dElapsed_1h_ms - CONST_DTICK_1H;
   
   	OUT_xOs_1h := 1;
   
   	IF NOT(OUT_xClock_1h) THEN
   		OUT_xClock_1h := 1;
   	ELSE
   		OUT_xClock_1h := 0;
   	END_IF;
   END_IF;
END_ROUTINE
END_ADD_ON_INSTRUCTION
